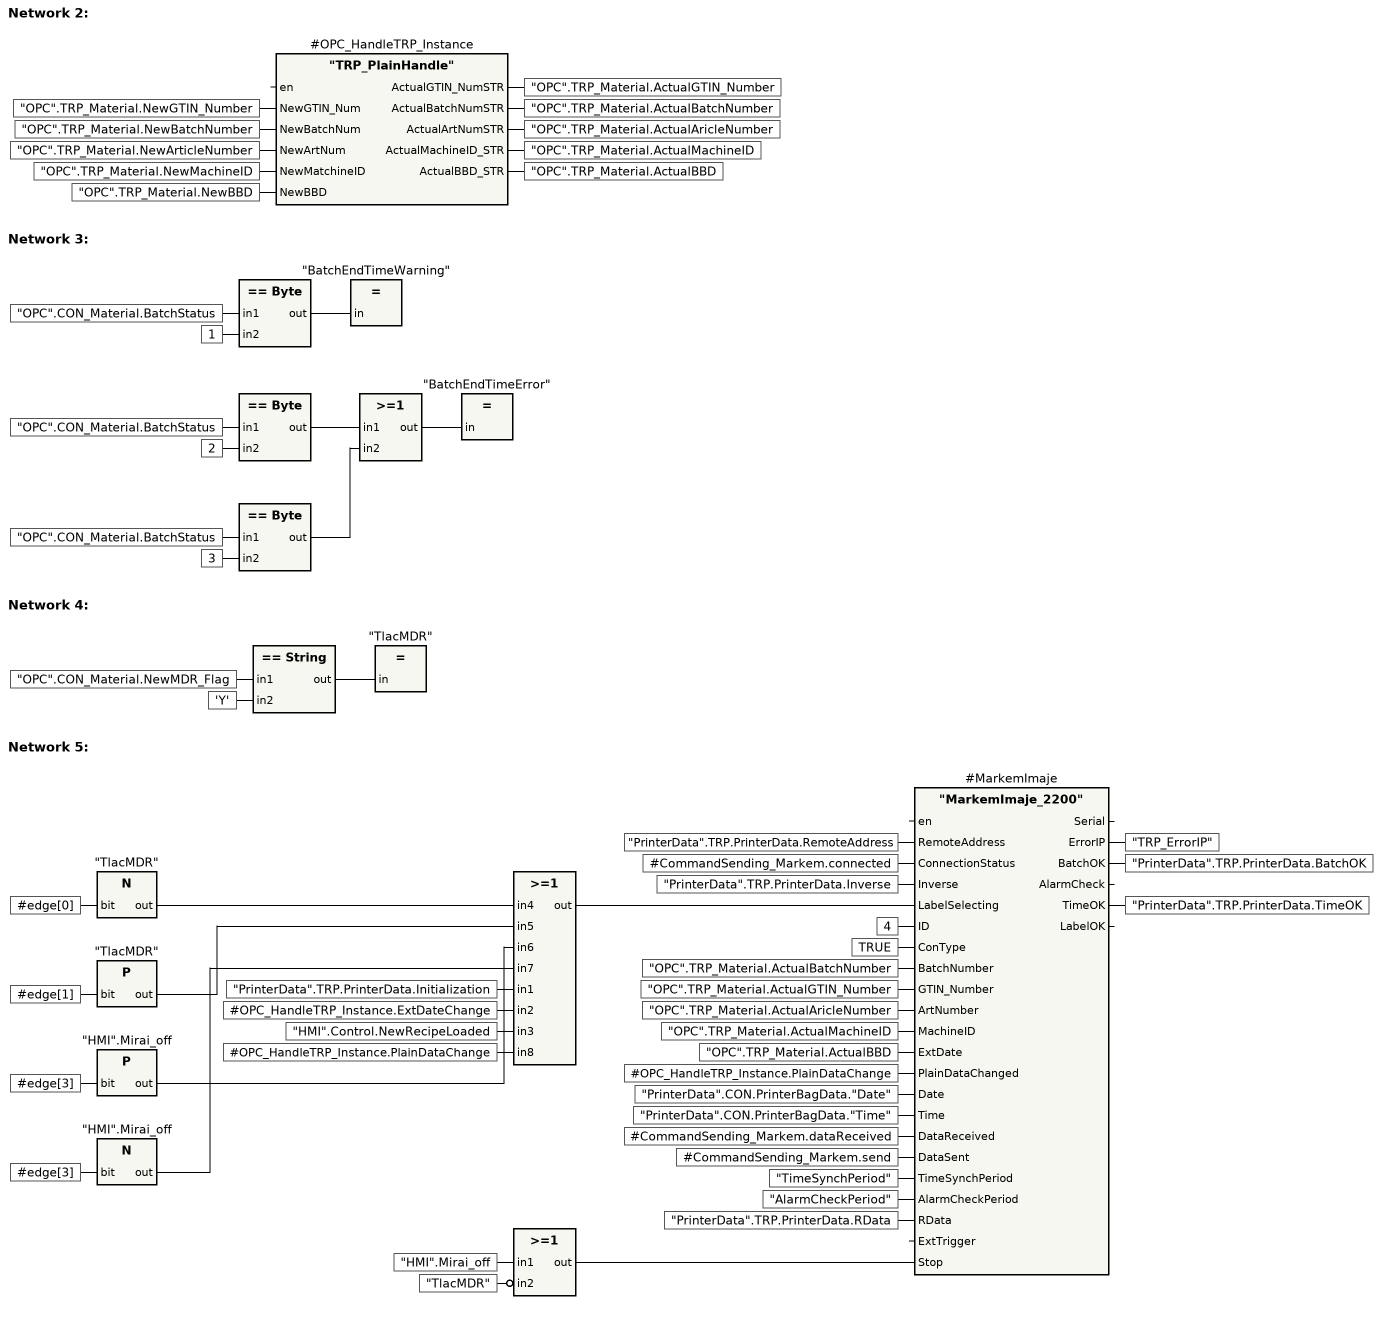
   #OPC_HandleTRP_Instance(NewGTIN_Num := "OPC".TRP_Material.NewGTIN_Number,   // "TRP_PlainHandle"
                           NewBatchNum := "OPC".TRP_Material.NewBatchNumber,
                           NewArtNum := "OPC".TRP_Material.NewArticleNumber,
                           NewMatchineID := "OPC".TRP_Material.NewMachineID,
                           NewBBD := "OPC".TRP_Material.NewBBD,
                           ActualGTIN_NumSTR => "OPC".TRP_Material.ActualGTIN_Number,
                           ActualBatchNumSTR => "OPC".TRP_Material.ActualBatchNumber,
                           ActualArtNumSTR => "OPC".TRP_Material.ActualAricleNumber,
                           ActualMachineID_STR => "OPC".TRP_Material.ActualMachineID,
                           ActualBBD_STR => "OPC".TRP_Material.ActualBBD);
END_REGION

REGION Network 3
   "BatchEndTimeWarning" := "OPC".CON_Material.BatchStatus = 1;
   "BatchEndTimeError" := ("OPC".CON_Material.BatchStatus = 2) OR ("OPC".CON_Material.BatchStatus = 3);
END_REGION

REGION Network 4
   // Porovnanie pre etiketovacku
   "TlacMDR" := "OPC".CON_Material.NewMDR_Flag = 'Y';
END_REGION

REGION Network 5
   #_w1 := NOT "TlacMDR" AND #edge[0];   // falling edge of "TlacMDR"
   #edge[0] := "TlacMDR";
   #_w2 := "TlacMDR" AND NOT #edge[1];   // rising edge of "TlacMDR"
   #edge[1] := "TlacMDR";
   #_w3 := "HMI".Mirai_off AND NOT #edge[3];   // rising edge of "HMI".Mirai_off
   #edge[3] := "HMI".Mirai_off;
   #_w4 := NOT "HMI".Mirai_off AND #edge[3];   // falling edge of "HMI".Mirai_off
   #edge[3] := "HMI".Mirai_off;
   #MarkemImaje(RemoteAddress := "PrinterData".TRP.PrinterData.RemoteAddress,   // "MarkemImaje_2200"
                ConnectionStatus := #CommandSending_Markem.connected,
                Inverse := "PrinterData".TRP.PrinterData.Inverse,
                LabelSelecting := #_w1 OR #_w2 OR #_w3 OR #_w4 OR "PrinterData".TRP.PrinterData.Initialization OR #OPC_HandleTRP_Instance.ExtDateChange OR "HMI".Control.NewRecipeLoaded OR #OPC_HandleTRP_Instance.PlainDataChange,
                ID := 4,
                ConType := TRUE,
                BatchNumber := "OPC".TRP_Material.ActualBatchNumber,
                GTIN_Number := "OPC".TRP_Material.ActualGTIN_Number,
                ArtNumber := "OPC".TRP_Material.ActualAricleNumber,
                MachineID := "OPC".TRP_Material.ActualMachineID,
                ExtDate := "OPC".TRP_Material.ActualBBD,
                PlainDataChanged := #OPC_HandleTRP_Instance.PlainDataChange,
                "Date" := "PrinterData".CON.PrinterBagData."Date",
                "Time" := "PrinterData".CON.PrinterBagData."Time",
                DataReceived := #CommandSending_Markem.dataReceived,
                DataSent := #CommandSending_Markem.send,
                TimeSynchPeriod := "TimeSynchPeriod",
                AlarmCheckPeriod := "AlarmCheckPeriod",
                RData := "PrinterData".TRP.PrinterData.RData,
                Stop := "HMI".Mirai_off OR NOT "TlacMDR",
                ErrorIP => "TRP_ErrorIP",
                BatchOK => "PrinterData".TRP.PrinterData.BatchOK,
                TimeOK => "PrinterData".TRP.PrinterData.TimeOK);
END_REGION

REGION Network 7
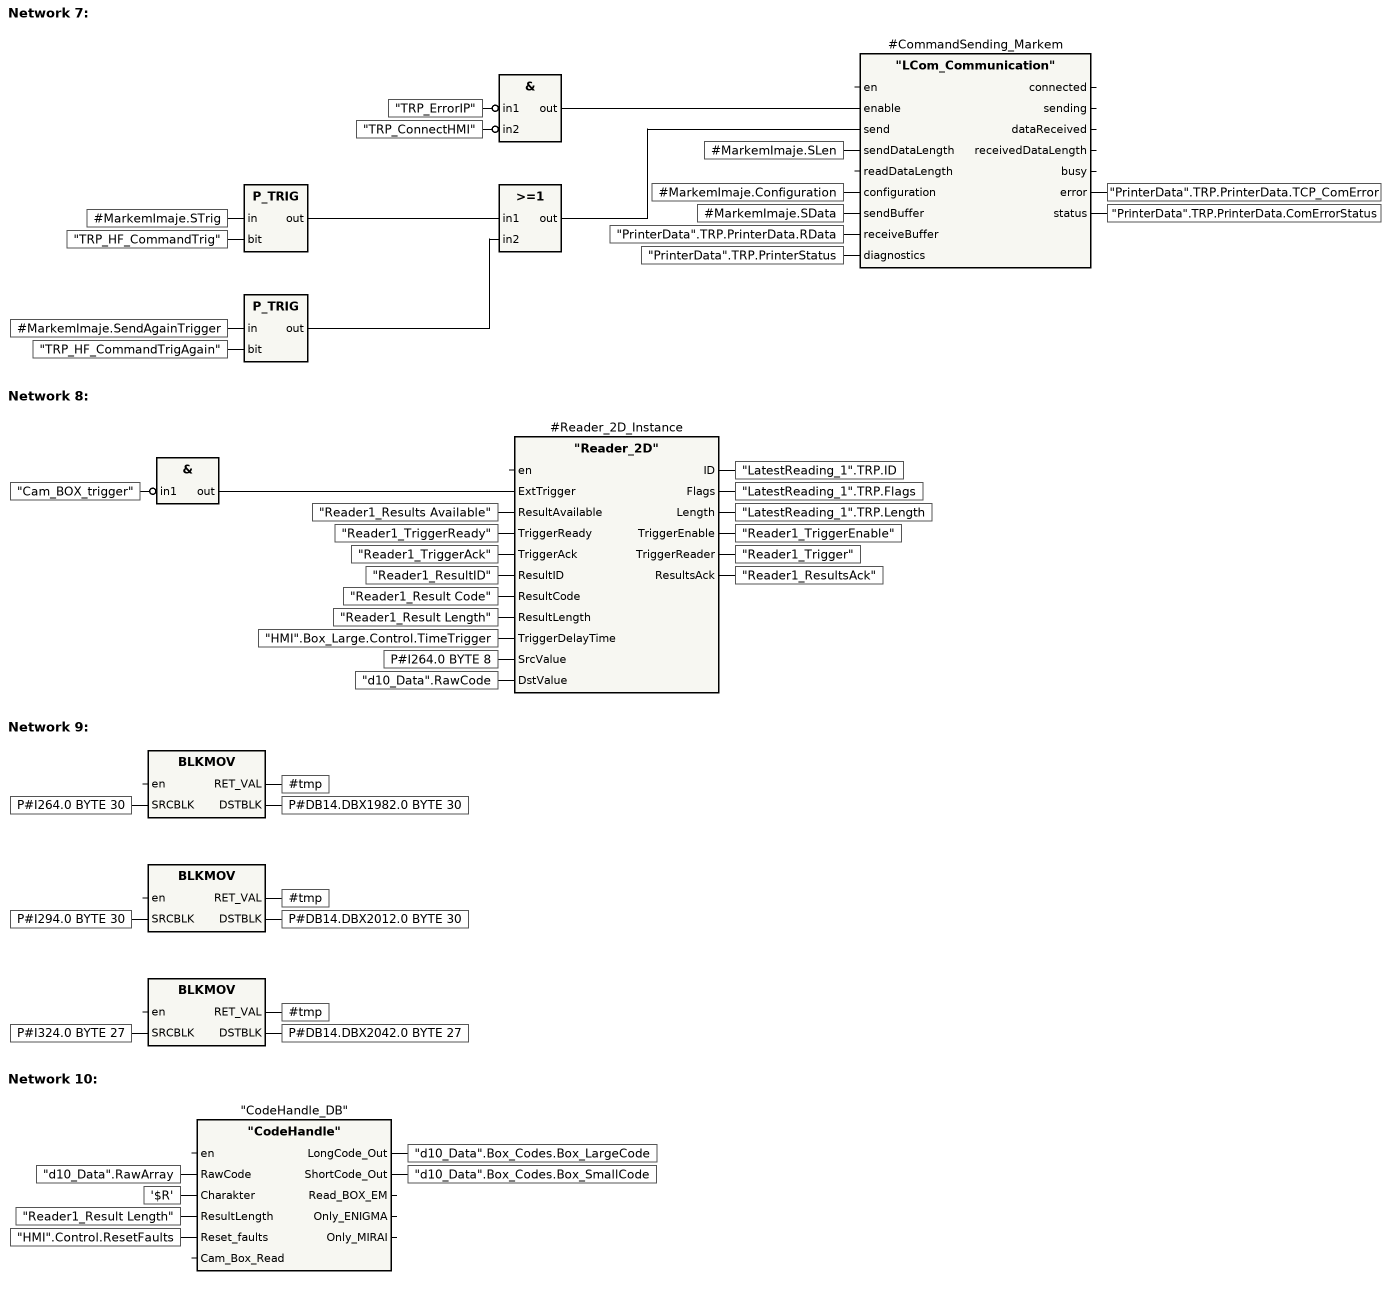
   #_w1 := #MarkemImaje.STrig AND NOT "TRP_HF_CommandTrig";   // rising edge
   "TRP_HF_CommandTrig" := #MarkemImaje.STrig;
   #_w2 := #MarkemImaje.SendAgainTrigger AND NOT "TRP_HF_CommandTrigAgain";   // rising edge
   "TRP_HF_CommandTrigAgain" := #MarkemImaje.SendAgainTrigger;
   #CommandSending_Markem(enable := NOT "TRP_ErrorIP" AND NOT "TRP_ConnectHMI",   // "LCom_Communication"
                          send := #_w1 OR #_w2,
                          sendDataLength := #MarkemImaje.SLen,
                          configuration := #MarkemImaje.Configuration,
                          sendBuffer := #MarkemImaje.SData,
                          receiveBuffer := "PrinterData".TRP.PrinterData.RData,
                          diagnostics := "PrinterData".TRP.PrinterStatus,
                          error => "PrinterData".TRP.PrinterData.TCP_ComError,
                          status => "PrinterData".TRP.PrinterData.ComErrorStatus);
END_REGION

REGION Network 8
   #Reader_2D_Instance(ExtTrigger := NOT "Cam_BOX_trigger",   // "Reader_2D"
                       ResultAvailable := "Reader1_Results Available",
                       TriggerReady := "Reader1_TriggerReady",
                       TriggerAck := "Reader1_TriggerAck",
                       ResultID := "Reader1_ResultID",
                       ResultCode := "Reader1_Result Code",
                       ResultLength := "Reader1_Result Length",
                       TriggerDelayTime := "HMI".Box_Large.Control.TimeTrigger,
                       SrcValue := P#I264.0 BYTE 8,
                       DstValue := "d10_Data".RawCode,
                       ID => "LatestReading_1".TRP.ID,
                       Flags => "LatestReading_1".TRP.Flags,
                       Length => "LatestReading_1".TRP.Length,
                       TriggerEnable => "Reader1_TriggerEnable",
                       TriggerReader => "Reader1_Trigger",
                       ResultsAck => "Reader1_ResultsAck");
END_REGION

REGION Network 9
   #tmp := BLKMOV(SRCBLK := P#I264.0 BYTE 30, DSTBLK => P#DB14.DBX1982.0 BYTE 30);
   #tmp := BLKMOV(SRCBLK := P#I294.0 BYTE 30, DSTBLK => P#DB14.DBX2012.0 BYTE 30);
   #tmp := BLKMOV(SRCBLK := P#I324.0 BYTE 27, DSTBLK => P#DB14.DBX2042.0 BYTE 27);
END_REGION

REGION Network 10
   "CodeHandle_DB"(RawCode := "d10_Data".RawArray,   // "CodeHandle"
                   Charakter := '$R',
                   ResultLength := "Reader1_Result Length",
                   Reset_faults := "HMI".Control.ResetFaults,
                   LongCode_Out => "d10_Data".Box_Codes.Box_LargeCode,
                   ShortCode_Out => "d10_Data".Box_Codes.Box_SmallCode);
END_REGION

REGION Network 11
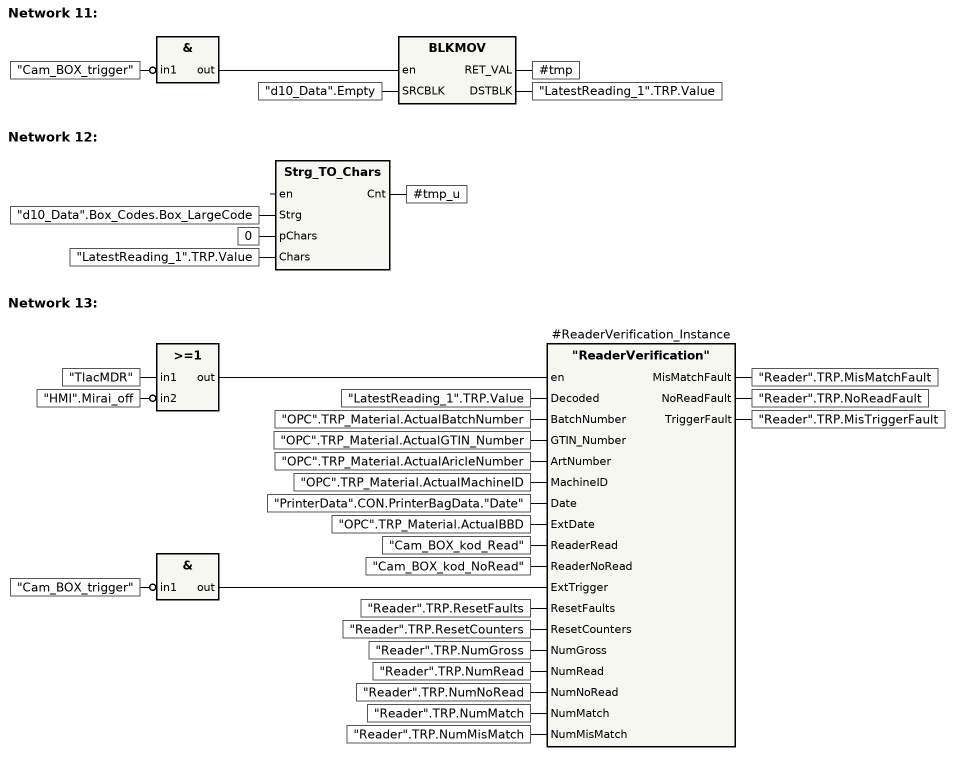
   IF NOT "Cam_BOX_trigger" THEN
       #tmp := BLKMOV(SRCBLK := "d10_Data".Empty, DSTBLK => "LatestReading_1".TRP.Value);
   END_IF;
END_REGION

REGION Network 12
   // no SCL statement known for Strg_TO_Chars: written as a call
   Strg_TO_Chars(Strg := "d10_Data".Box_Codes.Box_LargeCode,
                 pChars := 0,
                 Chars := "LatestReading_1".TRP.Value,
                 Cnt => #tmp_u);
END_REGION

REGION Network 13
   IF "TlacMDR" OR NOT "HMI".Mirai_off THEN
       #ReaderVerification_Instance(Decoded := "LatestReading_1".TRP.Value,   // "ReaderVerification"
                               BatchNumber := "OPC".TRP_Material.ActualBatchNumber,
                               GTIN_Number := "OPC".TRP_Material.ActualGTIN_Number,
                               ArtNumber := "OPC".TRP_Material.ActualAricleNumber,
                               MachineID := "OPC".TRP_Material.ActualMachineID,
                               "Date" := "PrinterData".CON.PrinterBagData."Date",
                               ExtDate := "OPC".TRP_Material.ActualBBD,
                               ReaderRead := "Cam_BOX_kod_Read",
                               ReaderNoRead := "Cam_BOX_kod_NoRead",
                               ExtTrigger := NOT "Cam_BOX_trigger",
                               ResetFaults := "Reader".TRP.ResetFaults,
                               ResetCounters := "Reader".TRP.ResetCounters,
                               NumGross := "Reader".TRP.NumGross,
                               NumRead := "Reader".TRP.NumRead,
                               NumNoRead := "Reader".TRP.NumNoRead,
                               NumMatch := "Reader".TRP.NumMatch,
                               NumMisMatch := "Reader".TRP.NumMisMatch,
                               MisMatchFault => "Reader".TRP.MisMatchFault,
                               NoReadFault => "Reader".TRP.NoReadFault,
                               TriggerFault => "Reader".TRP.MisTriggerFault);
   END_IF;
END_REGION

REGION Network 14
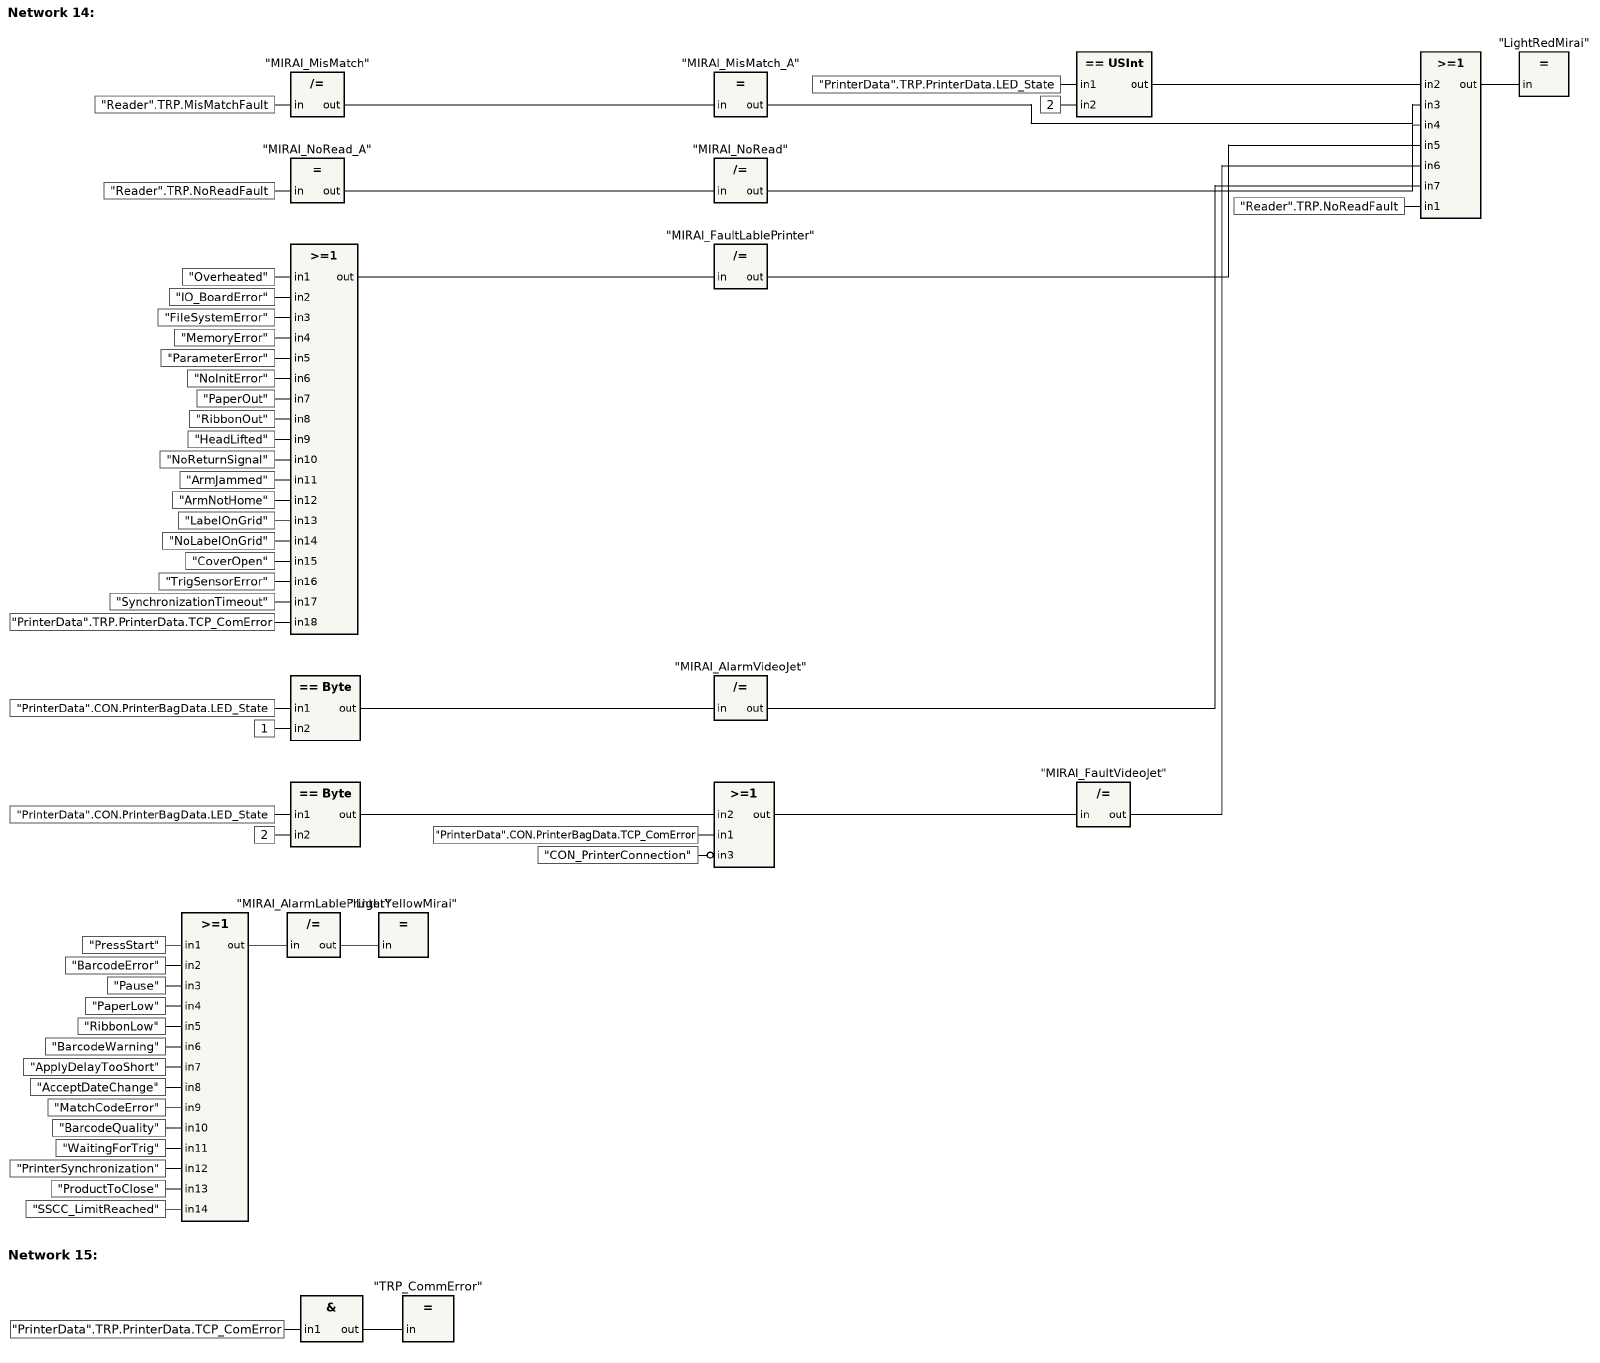
   "MIRAI_MisMatch" := NOT "Reader".TRP.MisMatchFault;
   "MIRAI_MisMatch_A" := "Reader".TRP.MisMatchFault;
   "MIRAI_NoRead_A" := "Reader".TRP.NoReadFault;
   "MIRAI_NoRead" := NOT "Reader".TRP.NoReadFault;
   #_w1 := "Overheated" OR "IO_BoardError" OR "FileSystemError" OR "MemoryError" OR "ParameterError" OR "NoInitError" OR "PaperOut" OR "RibbonOut" OR "HeadLifted" OR "NoReturnSignal" OR "ArmJammed" OR "ArmNotHome" OR "LabelOnGrid" OR "NoLabelOnGrid" OR "CoverOpen" OR "TrigSensorError" OR "SynchronizationTimeout" OR "PrinterData".TRP.PrinterData.TCP_ComError;
   "MIRAI_FaultLablePrinter" := NOT #_w1;
   #_w2 := ("PrinterData".CON.PrinterBagData.LED_State = 2) OR "PrinterData".CON.PrinterBagData.TCP_ComError OR NOT "CON_PrinterConnection";
   "MIRAI_FaultVideoJet" := NOT #_w2;
   #_w3 := "PrinterData".CON.PrinterBagData.LED_State = 1;
   "MIRAI_AlarmVideoJet" := NOT #_w3;
   "LightRedMirai" := ("PrinterData".TRP.PrinterData.LED_State = 2) OR "Reader".TRP.MisMatchFault OR "Reader".TRP.NoReadFault OR #_w1 OR #_w2 OR #_w3 OR "Reader".TRP.NoReadFault;
   #_w4 := "PressStart" OR "BarcodeError" OR "Pause" OR "PaperLow" OR "RibbonLow" OR "BarcodeWarning" OR "ApplyDelayTooShort" OR "AcceptDateChange" OR "MatchCodeError" OR "BarcodeQuality" OR "WaitingForTrig" OR "PrinterSynchronization" OR "ProductToClose" OR "SSCC_LimitReached";
   "MIRAI_AlarmLablePrinter" := NOT #_w4;
   "LightYellowMirai" := #_w4;
END_REGION

REGION Network 15
   "TRP_CommError" := "PrinterData".TRP.PrinterData.TCP_ComError;
END_REGION

REGION Network 16
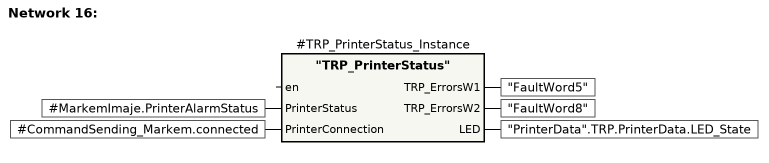
   #TRP_PrinterStatus_Instance(PrinterStatus := #MarkemImaje.PrinterAlarmStatus,   // "TRP_PrinterStatus"
                           PrinterConnection := #CommandSending_Markem.connected,
                           TRP_ErrorsW1 => "FaultWord5",
                           TRP_ErrorsW2 => "FaultWord8",
                           LED => "PrinterData".TRP.PrinterData.LED_State);
END_REGION
END_FUNCTION_BLOCK

FUNCTION_BLOCK "ProgramReaderBox"   // FB11, FBD
{ S7_Optimized_Access := 'TRUE' }
VERSION : 0.1
   VAR
      HandleCom_Instance : "HandleCom";
      SimpleRead_Instance : "SimpleRead";
      ProgramReader_Instance : "ProgramReader";
      IEC_Timer_0_Instance : TON_TIME;
      t_DelayNoRead : TON_TIME;
   END_VAR
   VAR_TEMP
      TmpW : Word;
   END_VAR
BEGIN

REGION Network 1
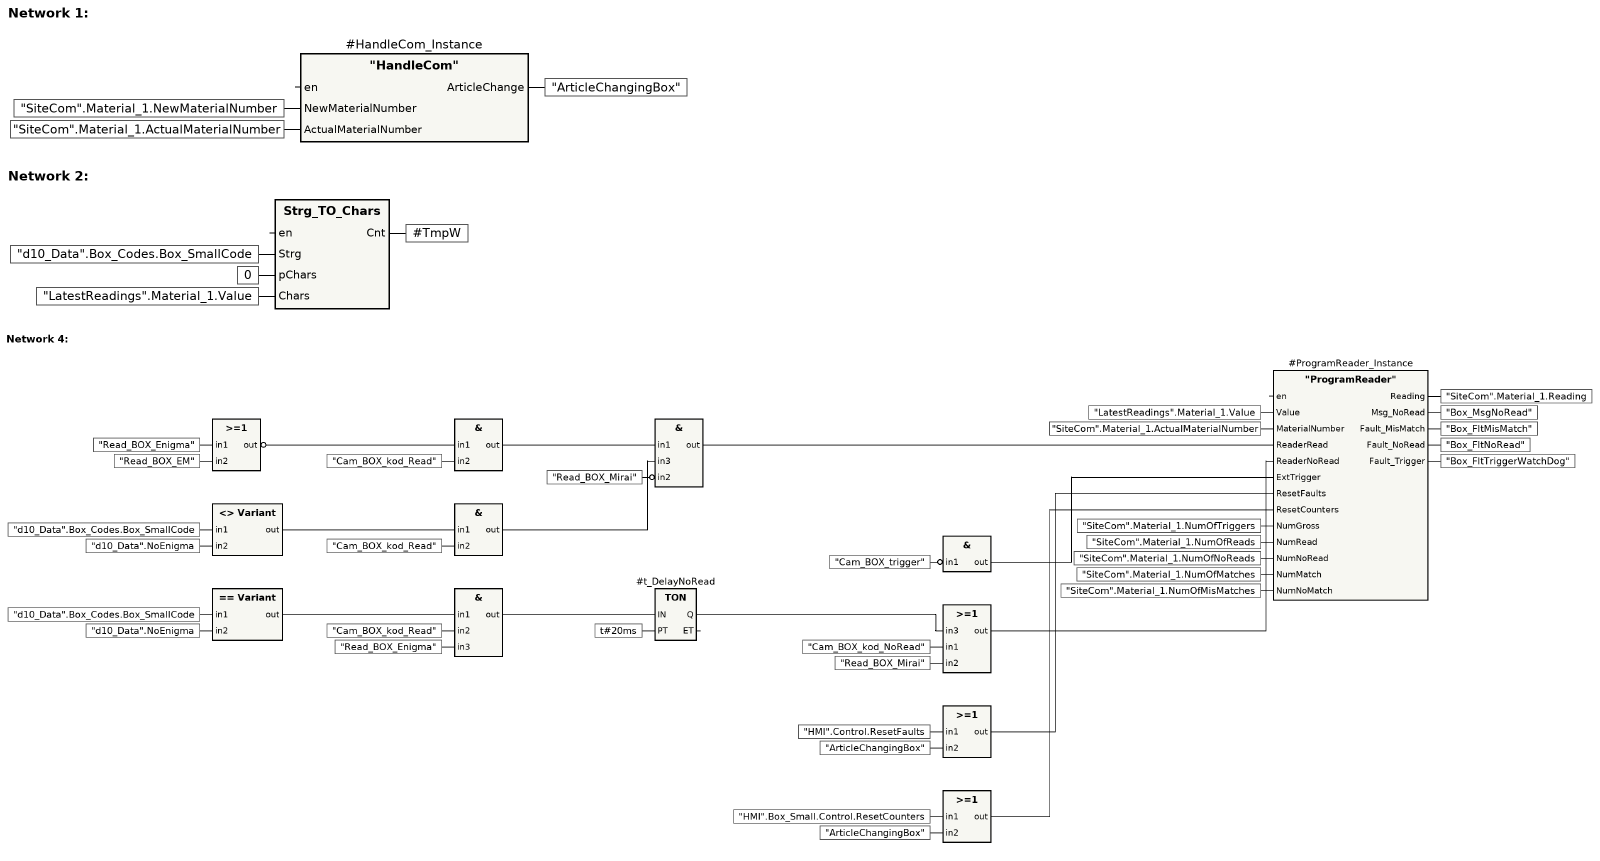
   #HandleCom_Instance(NewMaterialNumber := "SiteCom".Material_1.NewMaterialNumber,   // "HandleCom"
                       ActualMaterialNumber := "SiteCom".Material_1.ActualMaterialNumber,
                       ArticleChange => "ArticleChangingBox");
END_REGION

REGION Network 2
   // no SCL statement known for Strg_TO_Chars: written as a call
   Strg_TO_Chars(Strg := "d10_Data".Box_Codes.Box_SmallCode,
                 pChars := 0,
                 Chars := "LatestReadings".Material_1.Value,
                 Cnt => #TmpW);
END_REGION

REGION Network 4
   #t_DelayNoRead(IN := ("d10_Data".Box_Codes.Box_SmallCode = "d10_Data".NoEnigma) AND "Cam_BOX_kod_Read" AND "Read_BOX_Enigma",   // TON
                  PT := t#20ms);
   #ProgramReader_Instance(Value := "LatestReadings".Material_1.Value,   // "ProgramReader"
                           MaterialNumber := "SiteCom".Material_1.ActualMaterialNumber,
                           ReaderRead := NOT ("Read_BOX_Enigma" OR "Read_BOX_EM") AND "Cam_BOX_kod_Read" AND ("d10_Data".Box_Codes.Box_SmallCode <> "d10_Data".NoEnigma) AND "Cam_BOX_kod_Read" AND NOT "Read_BOX_Mirai",
                           ReaderNoRead := #t_DelayNoRead.Q OR "Cam_BOX_kod_NoRead" OR "Read_BOX_Mirai",
                           ExtTrigger := NOT "Cam_BOX_trigger",
                           ResetFaults := "HMI".Control.ResetFaults OR "ArticleChangingBox",
                           ResetCounters := "HMI".Box_Small.Control.ResetCounters OR "ArticleChangingBox",
                           NumGross := "SiteCom".Material_1.NumOfTriggers,
                           NumRead := "SiteCom".Material_1.NumOfReads,
                           NumNoRead := "SiteCom".Material_1.NumOfNoReads,
                           NumMatch := "SiteCom".Material_1.NumOfMatches,
                           NumNoMatch := "SiteCom".Material_1.NumOfMisMatches,
                           Reading => "SiteCom".Material_1.Reading,
                           Msg_NoRead => "Box_MsgNoRead",
                           Fault_MisMatch => "Box_FltMisMatch",
                           Fault_NoRead => "Box_FltNoRead",
                           Fault_Trigger => "Box_FltTriggerWatchDog");
END_REGION

REGION Network 5
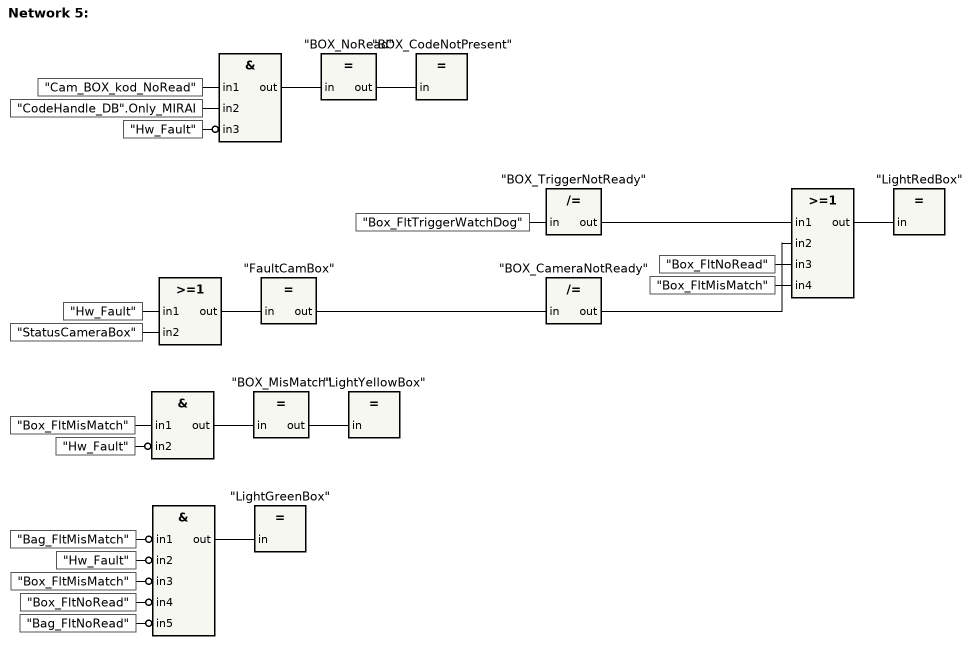
   "BOX_NoRead" := "Cam_BOX_kod_NoRead" AND "CodeHandle_DB".Only_MIRAI AND NOT "Hw_Fault";
   "BOX_CodeNotPresent" := "BOX_NoRead";
   "BOX_TriggerNotReady" := NOT "Box_FltTriggerWatchDog";
   "FaultCamBox" := "Hw_Fault" OR "StatusCameraBox";
   "BOX_CameraNotReady" := NOT "FaultCamBox";
   "LightRedBox" := "Box_FltTriggerWatchDog" OR "FaultCamBox" OR "Box_FltNoRead" OR "Box_FltMisMatch";
   "BOX_MisMatch" := "Box_FltMisMatch" AND NOT "Hw_Fault";
   "LightYellowBox" := "BOX_MisMatch";
   "LightGreenBox" := NOT "Bag_FltMisMatch" AND NOT "Hw_Fault" AND NOT "Box_FltMisMatch" AND NOT "Box_FltNoRead" AND NOT "Bag_FltNoRead";
END_REGION
END_FUNCTION_BLOCK

FUNCTION_BLOCK "ProgramReaderBag"   // FB12, FBD
{ S7_Optimized_Access := 'TRUE' }
VERSION : 0.1
   VAR
      HandleCom_Instance : "HandleCom";
      SimpleRead_Instance : "SimpleRead";
      ProgramReader_Instance : "ProgramReader";
      IEC_Timer_0_Instance : TON_TIME;
   END_VAR
BEGIN

REGION Network 2
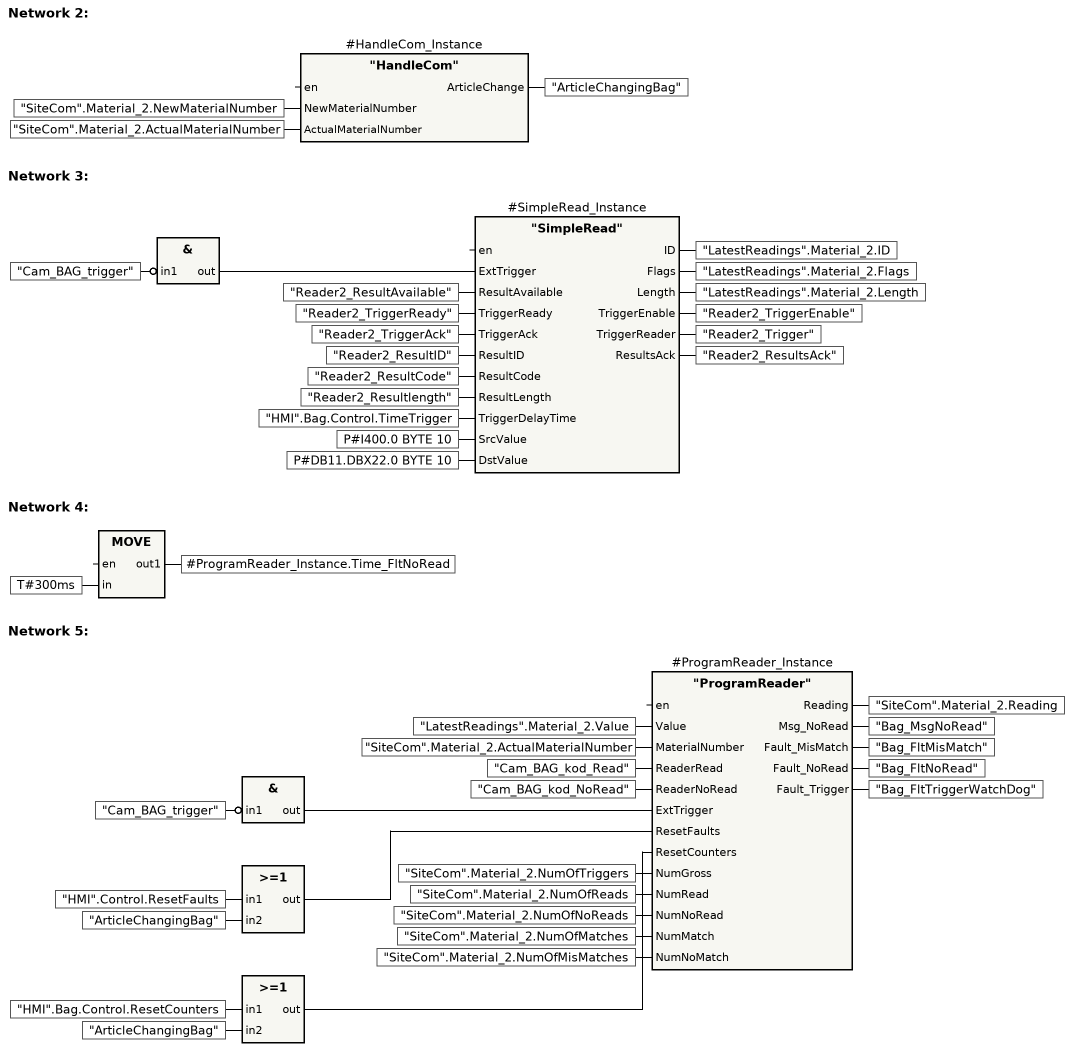
   #HandleCom_Instance(NewMaterialNumber := "SiteCom".Material_2.NewMaterialNumber,   // "HandleCom"
                       ActualMaterialNumber := "SiteCom".Material_2.ActualMaterialNumber,
                       ArticleChange => "ArticleChangingBag");
END_REGION

REGION Network 3
   #SimpleRead_Instance(ExtTrigger := NOT "Cam_BAG_trigger",   // "SimpleRead"
                        ResultAvailable := "Reader2_ResultAvailable",
                        TriggerReady := "Reader2_TriggerReady",
                        TriggerAck := "Reader2_TriggerAck",
                        ResultID := "Reader2_ResultID",
                        ResultCode := "Reader2_ResultCode",
                        ResultLength := "Reader2_Resultlength",
                        TriggerDelayTime := "HMI".Bag.Control.TimeTrigger,
                        SrcValue := P#I400.0 BYTE 10,
                        DstValue := P#DB11.DBX22.0 BYTE 10,
                        ID => "LatestReadings".Material_2.ID,
                        Flags => "LatestReadings".Material_2.Flags,
                        Length => "LatestReadings".Material_2.Length,
                        TriggerEnable => "Reader2_TriggerEnable",
                        TriggerReader => "Reader2_Trigger",
                        ResultsAck => "Reader2_ResultsAck");
END_REGION

REGION Network 4
   #ProgramReader_Instance.Time_FltNoRead := T#300ms;
END_REGION

REGION Network 5
   #ProgramReader_Instance(Value := "LatestReadings".Material_2.Value,   // "ProgramReader"
                           MaterialNumber := "SiteCom".Material_2.ActualMaterialNumber,
                           ReaderRead := "Cam_BAG_kod_Read",
                           ReaderNoRead := "Cam_BAG_kod_NoRead",
                           ExtTrigger := NOT "Cam_BAG_trigger",
                           ResetFaults := "HMI".Control.ResetFaults OR "ArticleChangingBag",
                           ResetCounters := "HMI".Bag.Control.ResetCounters OR "ArticleChangingBag",
                           NumGross := "SiteCom".Material_2.NumOfTriggers,
                           NumRead := "SiteCom".Material_2.NumOfReads,
                           NumNoRead := "SiteCom".Material_2.NumOfNoReads,
                           NumMatch := "SiteCom".Material_2.NumOfMatches,
                           NumNoMatch := "SiteCom".Material_2.NumOfMisMatches,
                           Reading => "SiteCom".Material_2.Reading,
                           Msg_NoRead => "Bag_MsgNoRead",
                           Fault_MisMatch => "Bag_FltMisMatch",
                           Fault_NoRead => "Bag_FltNoRead",
                           Fault_Trigger => "Bag_FltTriggerWatchDog");
END_REGION

REGION Network 6
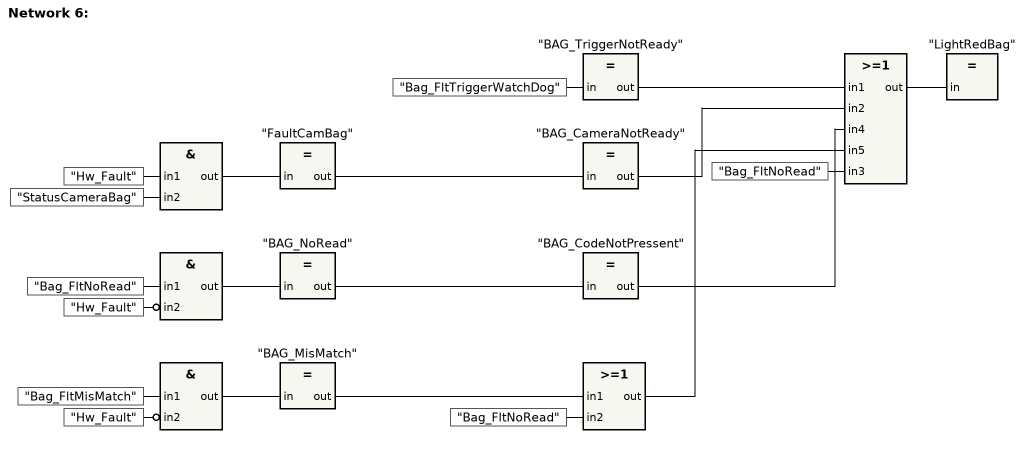
   "BAG_TriggerNotReady" := "Bag_FltTriggerWatchDog";
   "FaultCamBag" := "Hw_Fault" AND "StatusCameraBag";
   "BAG_CameraNotReady" := "FaultCamBag";
   "BAG_NoRead" := "Bag_FltNoRead" AND NOT "Hw_Fault";
   "BAG_CodeNotPressent" := "BAG_NoRead";
   "BAG_MisMatch" := "Bag_FltMisMatch" AND NOT "Hw_Fault";
   "LightRedBag" := "Bag_FltTriggerWatchDog" OR "FaultCamBag" OR "BAG_NoRead" OR "BAG_MisMatch" OR "Bag_FltNoRead" OR "Bag_FltNoRead";
END_REGION
END_FUNCTION_BLOCK

FUNCTION_BLOCK "CON"   // FB13, FBD
{ S7_Optimized_Access := 'TRUE' }
VERSION : 0.1
   VAR
      HandleComBag : "CON_PlainHandle";
      Domino : "Domino_AX";
      ComandsSending_Domino : "LCom_Communication";
      BatchSending_Domino : "LCom_Communication";
      VideoJet : "VideoJet_1520";
      ComandsSending_Video : "LCom_Communication";
      CON_PrinterStatus_Instance : "CON_PrinterStatus";
   END_VAR
   VAR_TEMP   // added for the SCL form of the ladder/FBD networks
      _w1 : Bool;
      _w2 : Bool;
   END_VAR
BEGIN

REGION Network 1
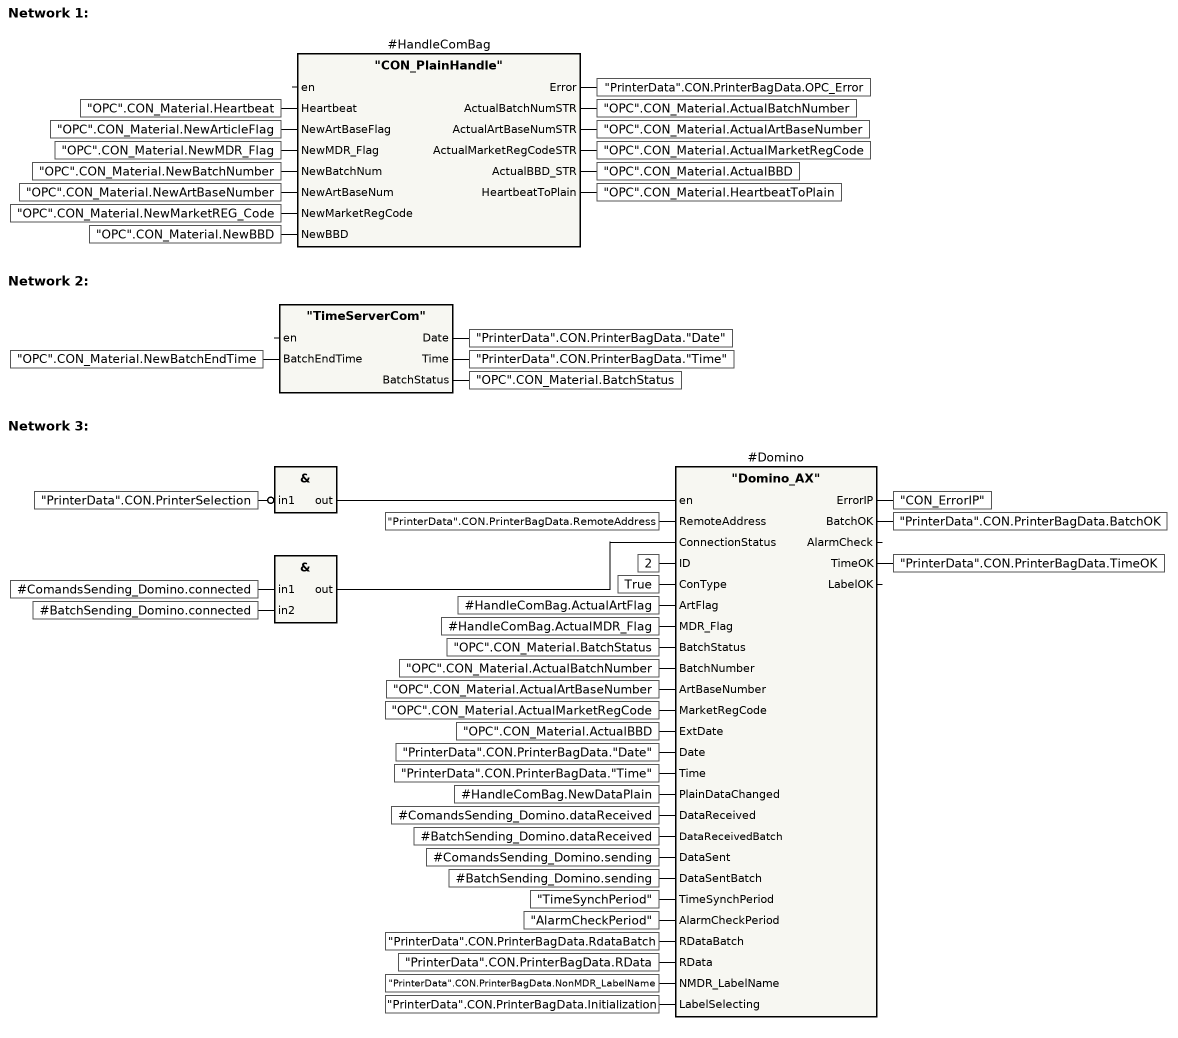
   #HandleComBag(Heartbeat := "OPC".CON_Material.Heartbeat,   // "CON_PlainHandle"
                 NewArtBaseFlag := "OPC".CON_Material.NewArticleFlag,
                 NewMDR_Flag := "OPC".CON_Material.NewMDR_Flag,
                 NewBatchNum := "OPC".CON_Material.NewBatchNumber,
                 NewArtBaseNum := "OPC".CON_Material.NewArtBaseNumber,
                 NewMarketRegCode := "OPC".CON_Material.NewMarketREG_Code,
                 NewBBD := "OPC".CON_Material.NewBBD,
                 Error => "PrinterData".CON.PrinterBagData.OPC_Error,
                 ActualBatchNumSTR => "OPC".CON_Material.ActualBatchNumber,
                 ActualArtBaseNumSTR => "OPC".CON_Material.ActualArtBaseNumber,
                 ActualMarketRegCodeSTR => "OPC".CON_Material.ActualMarketRegCode,
                 ActualBBD_STR => "OPC".CON_Material.ActualBBD,
                 HeartbeatToPlain => "OPC".CON_Material.HeartbeatToPlain);
END_REGION
